// TIA Portal project "SMSS-ENLAB-01-003-1508-012-PLC-B_V13_SP1_1_V17" (V17) (continued)
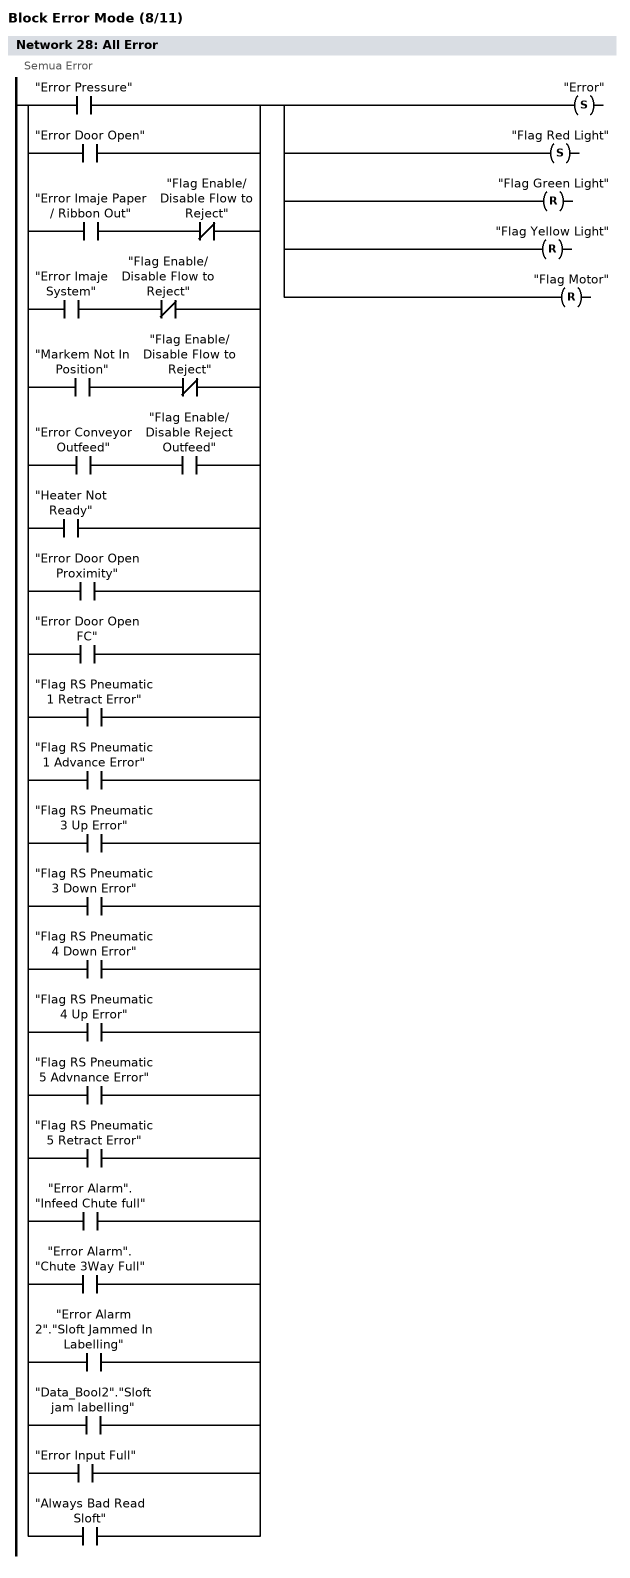
   RUNG wire#powerrail
      Contact( "Error Pressure" )
      wire#w1
      S_Coil( "Error" )
   END_RUNG
   RUNG wire#powerrail
      Contact( "Error Door Open" )
   END_RUNG wire#w1
   RUNG wire#powerrail
      Contact( "Error Imaje Paper / Ribbon Out" )
      I_Contact( "Flag Enable/Disable Flow to Reject" )
   END_RUNG wire#w1
   RUNG wire#powerrail
      Contact( "Error Imaje System" )
      I_Contact( "Flag Enable/Disable Flow to Reject" )
   END_RUNG wire#w1
   RUNG wire#powerrail
      Contact( "Markem Not In Position" )
      I_Contact( "Flag Enable/Disable Flow to Reject" )
   END_RUNG wire#w1
   RUNG wire#powerrail
      Contact( "Error Conveyor Outfeed" )
      Contact( "Flag Enable/Disable Reject Outfeed" )
   END_RUNG wire#w1
   RUNG wire#powerrail
      Contact( "Heater Not Ready" )
   END_RUNG wire#w1
   RUNG wire#powerrail
      Contact( "Error Door Open Proximity" )
   END_RUNG wire#w1
   RUNG wire#powerrail
      Contact( "Error Door Open FC" )
   END_RUNG wire#w1
   RUNG wire#powerrail
      Contact( "Flag RS Pneumatic 1 Retract Error" )
   END_RUNG wire#w1
   RUNG wire#powerrail
      Contact( "Flag RS Pneumatic 1 Advance Error" )
   END_RUNG wire#w1
   RUNG wire#powerrail
      Contact( "Flag RS Pneumatic 3 Up Error" )
   END_RUNG wire#w1
   RUNG wire#powerrail
      Contact( "Flag RS Pneumatic 3 Down Error" )
   END_RUNG wire#w1
   RUNG wire#powerrail
      Contact( "Flag RS Pneumatic 4 Down Error" )
   END_RUNG wire#w1
   RUNG wire#powerrail
      Contact( "Flag RS Pneumatic 4 Up Error" )
   END_RUNG wire#w1
   RUNG wire#powerrail
      Contact( "Flag RS Pneumatic 5 Advnance Error" )
   END_RUNG wire#w1
   RUNG wire#powerrail
      Contact( "Flag RS Pneumatic 5 Retract Error" )
   END_RUNG wire#w1
   RUNG wire#powerrail
      Contact( "Error Alarm"."Infeed Chute full" )
   END_RUNG wire#w1
   RUNG wire#powerrail
      Contact( "Error Alarm"."Chute 3Way Full" )
   END_RUNG wire#w1
   RUNG wire#powerrail
      Contact( "Error Alarm 2"."Sloft Jammed In Labelling" )
   END_RUNG wire#w1
   RUNG wire#powerrail
      Contact( "Data_Bool2"."Sloft jam labelling" )
   END_RUNG wire#w1
   RUNG wire#powerrail
      Contact( "Error Input Full" )
   END_RUNG wire#w1
   RUNG wire#powerrail
      Contact( "Always Bad Read Sloft" )
   END_RUNG wire#w1
   RUNG wire#w1
      S_Coil( "Flag Red Light" )
   END_RUNG
   RUNG wire#w1
      R_Coil( "Flag Green Light" )
   END_RUNG
   RUNG wire#w1
      R_Coil( "Flag Yellow Light" )
   END_RUNG
   RUNG wire#w1
      R_Coil( "Flag Motor" )
   END_RUNG
   // the same network as SCL:
   IF "Error Pressure" OR "Error Door Open" OR ("Error Imaje Paper / Ribbon Out" AND NOT "Flag Enable/Disable Flow to Reject") OR ("Error Imaje System" AND NOT "Flag Enable/Disable Flow to Reject") OR ("Markem Not In Position" AND NOT "Flag Enable/Disable Flow to Reject") OR ("Error Conveyor Outfeed" AND "Flag Enable/Disable Reject Outfeed") OR "Heater Not Ready" OR "Error Door Open Proximity" OR "Error Door Open FC" OR "Flag RS Pneumatic 1 Retract Error" OR "Flag RS Pneumatic 1 Advance Error" OR "Flag RS Pneumatic 3 Up Error" OR "Flag RS Pneumatic 3 Down Error" OR "Flag RS Pneumatic 4 Down Error" OR "Flag RS Pneumatic 4 Up Error" OR "Flag RS Pneumatic 5 Advnance Error" OR "Flag RS Pneumatic 5 Retract Error" OR "Error Alarm"."Infeed Chute full" OR "Error Alarm"."Chute 3Way Full" OR "Error Alarm 2"."Sloft Jammed In Labelling" OR "Data_Bool2"."Sloft jam labelling" OR "Error Input Full" OR "Always Bad Read Sloft" THEN
       "Error" := TRUE;
       "Flag Red Light" := TRUE;
       "Flag Green Light" := FALSE;
       "Flag Yellow Light" := FALSE;
       "Flag Motor" := FALSE;
   END_IF;
END_REGION

REGION Network 29: Reset Error
   // Untuk Reset Semua Error
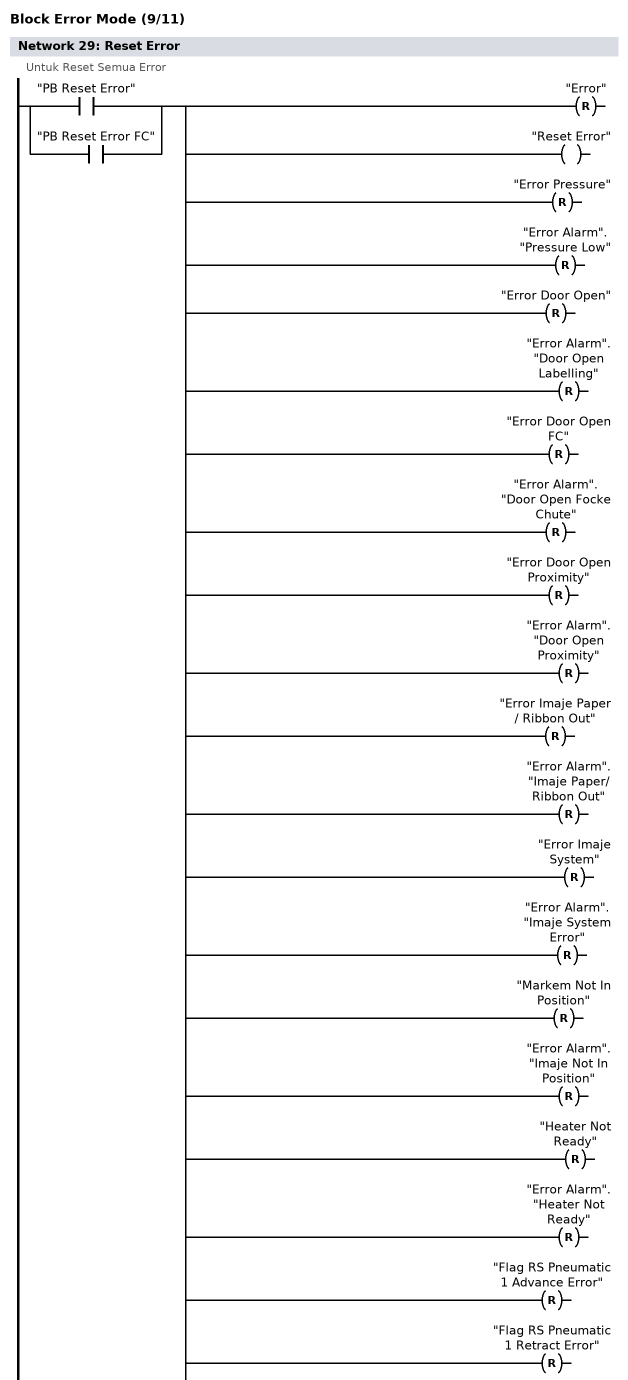
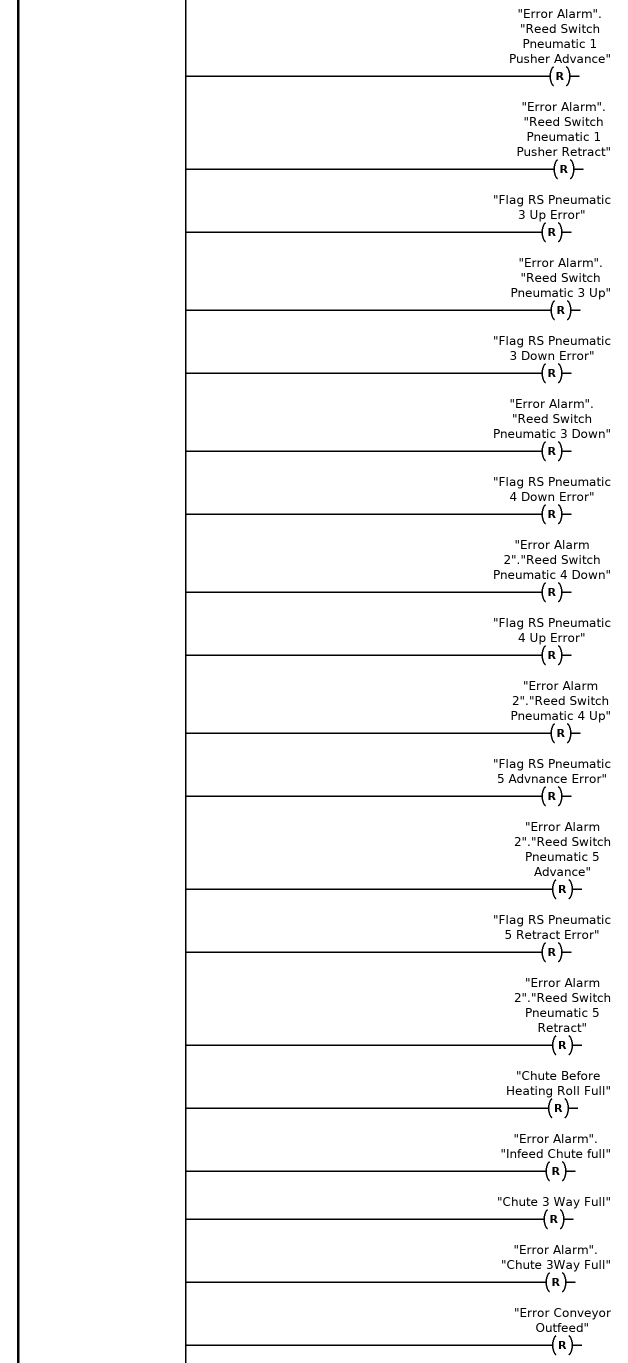
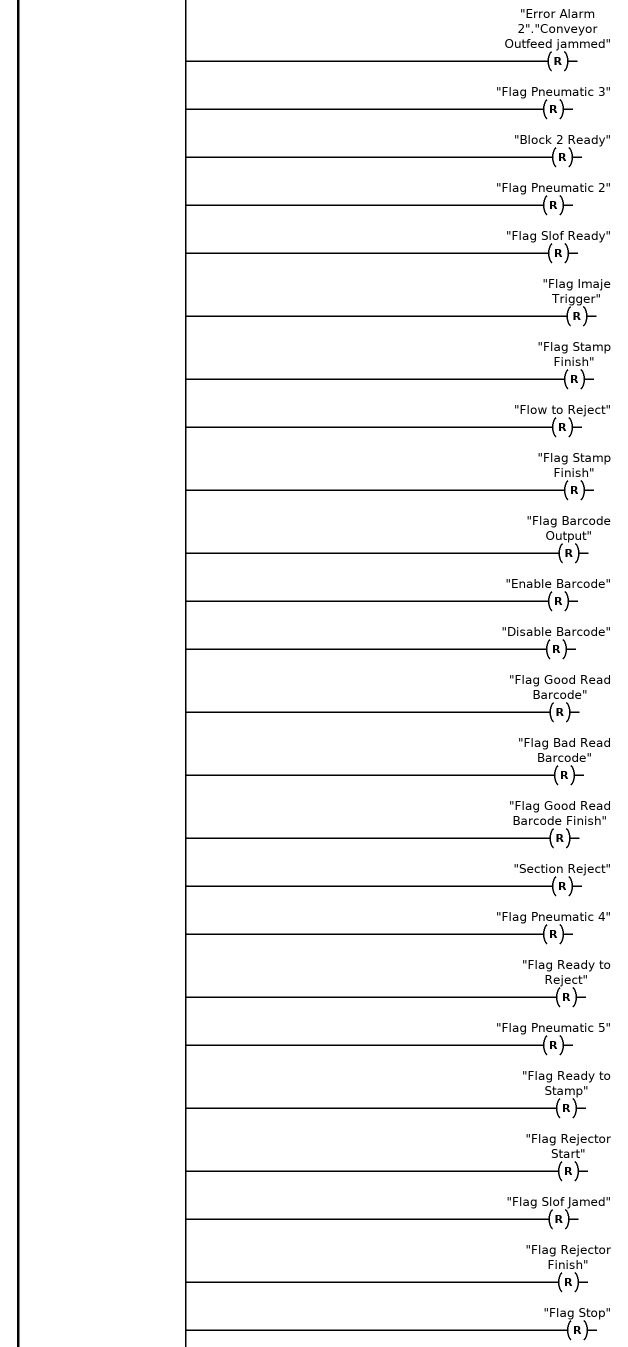
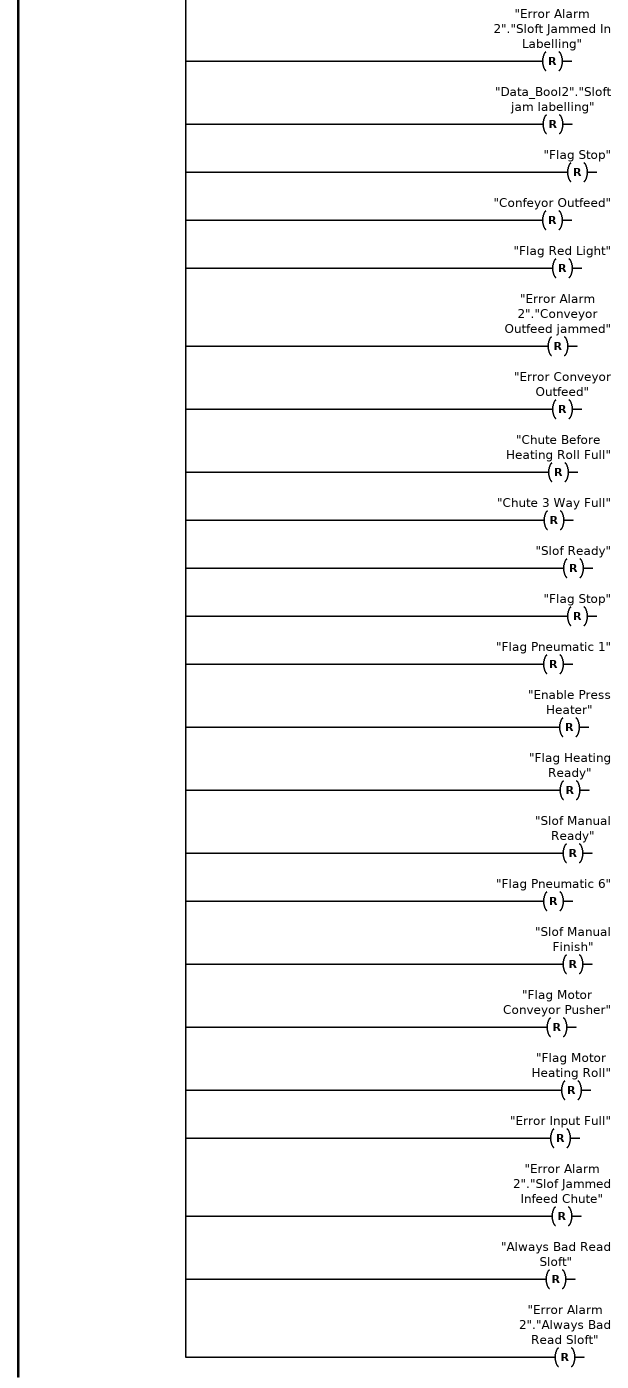
   RUNG wire#powerrail
      Contact( "PB Reset Error" )
      wire#w1
      R_Coil( "Error" )
   END_RUNG
   RUNG wire#powerrail
      Contact( "PB Reset Error FC" )
   END_RUNG wire#w1
   RUNG wire#w1
      Coil( "Reset Error" )
   END_RUNG
   RUNG wire#w1
      R_Coil( "Error Pressure" )
   END_RUNG
   RUNG wire#w1
      R_Coil( "Error Alarm"."Pressure Low" )
   END_RUNG
   RUNG wire#w1
      R_Coil( "Error Door Open" )
   END_RUNG
   RUNG wire#w1
      R_Coil( "Error Alarm"."Door Open Labelling" )
   END_RUNG
   RUNG wire#w1
      R_Coil( "Error Door Open FC" )
   END_RUNG
   RUNG wire#w1
      R_Coil( "Error Alarm"."Door Open Focke Chute" )
   END_RUNG
   RUNG wire#w1
      R_Coil( "Error Door Open Proximity" )
   END_RUNG
   RUNG wire#w1
      R_Coil( "Error Alarm"."Door Open Proximity" )
   END_RUNG
   RUNG wire#w1
      R_Coil( "Error Imaje Paper / Ribbon Out" )
   END_RUNG
   RUNG wire#w1
      R_Coil( "Error Alarm"."Imaje Paper/Ribbon Out" )
   END_RUNG
   RUNG wire#w1
      R_Coil( "Error Imaje System" )
   END_RUNG
   RUNG wire#w1
      R_Coil( "Error Alarm"."Imaje System Error" )
   END_RUNG
   RUNG wire#w1
      R_Coil( "Markem Not In Position" )
   END_RUNG
   RUNG wire#w1
      R_Coil( "Error Alarm"."Imaje Not In Position" )
   END_RUNG
   RUNG wire#w1
      R_Coil( "Heater Not Ready" )
   END_RUNG
   RUNG wire#w1
      R_Coil( "Error Alarm"."Heater Not Ready" )
   END_RUNG
   RUNG wire#w1
      R_Coil( "Flag RS Pneumatic 1 Advance Error" )
   END_RUNG
   RUNG wire#w1
      R_Coil( "Flag RS Pneumatic 1 Retract Error" )
   END_RUNG
   RUNG wire#w1
      R_Coil( "Error Alarm"."Reed Switch Pneumatic 1 Pusher Advance" )
   END_RUNG
   RUNG wire#w1
      R_Coil( "Error Alarm"."Reed Switch Pneumatic 1 Pusher Retract" )
   END_RUNG
   RUNG wire#w1
      R_Coil( "Flag RS Pneumatic 3 Up Error" )
   END_RUNG
   RUNG wire#w1
      R_Coil( "Error Alarm"."Reed Switch Pneumatic 3 Up" )
   END_RUNG
   RUNG wire#w1
      R_Coil( "Flag RS Pneumatic 3 Down Error" )
   END_RUNG
   RUNG wire#w1
      R_Coil( "Error Alarm"."Reed Switch Pneumatic 3 Down" )
   END_RUNG
   RUNG wire#w1
      R_Coil( "Flag RS Pneumatic 4 Down Error" )
   END_RUNG
   RUNG wire#w1
      R_Coil( "Error Alarm 2"."Reed Switch Pneumatic 4 Down" )
   END_RUNG
   RUNG wire#w1
      R_Coil( "Flag RS Pneumatic 4 Up Error" )
   END_RUNG
   RUNG wire#w1
      R_Coil( "Error Alarm 2"."Reed Switch Pneumatic 4 Up" )
   END_RUNG
   RUNG wire#w1
      R_Coil( "Flag RS Pneumatic 5 Advnance Error" )
   END_RUNG
   RUNG wire#w1
      R_Coil( "Error Alarm 2"."Reed Switch Pneumatic 5 Advance" )
   END_RUNG
   RUNG wire#w1
      R_Coil( "Flag RS Pneumatic 5 Retract Error" )
   END_RUNG
   RUNG wire#w1
      R_Coil( "Error Alarm 2"."Reed Switch Pneumatic 5 Retract" )
   END_RUNG
   RUNG wire#w1
      R_Coil( "Chute Before Heating Roll Full" )
   END_RUNG
   RUNG wire#w1
      R_Coil( "Error Alarm"."Infeed Chute full" )
   END_RUNG
   RUNG wire#w1
      R_Coil( "Chute 3 Way Full" )
   END_RUNG
   RUNG wire#w1
      R_Coil( "Error Alarm"."Chute 3Way Full" )
   END_RUNG
   RUNG wire#w1
      R_Coil( "Error Conveyor Outfeed" )
   END_RUNG
   RUNG wire#w1
      R_Coil( "Error Alarm 2"."Conveyor Outfeed jammed" )
   END_RUNG
   RUNG wire#w1
      R_Coil( "Flag Pneumatic 3" )
   END_RUNG
   RUNG wire#w1
      R_Coil( "Block 2 Ready" )
   END_RUNG
   RUNG wire#w1
      R_Coil( "Flag Pneumatic 2" )
   END_RUNG
   RUNG wire#w1
      R_Coil( "Flag Slof Ready" )
   END_RUNG
   RUNG wire#w1
      R_Coil( "Flag Imaje Trigger" )
   END_RUNG
   RUNG wire#w1
      R_Coil( "Flag Stamp Finish" )
   END_RUNG
   RUNG wire#w1
      R_Coil( "Flow to Reject" )
   END_RUNG
   RUNG wire#w1
      R_Coil( "Flag Stamp Finish" )
   END_RUNG
   RUNG wire#w1
      R_Coil( "Flag Barcode Output" )
   END_RUNG
   RUNG wire#w1
      R_Coil( "Enable Barcode" )
   END_RUNG
   RUNG wire#w1
      R_Coil( "Disable Barcode" )
   END_RUNG
   RUNG wire#w1
      R_Coil( "Flag Good Read Barcode" )
   END_RUNG
   RUNG wire#w1
      R_Coil( "Flag Bad Read Barcode" )
   END_RUNG
   RUNG wire#w1
      R_Coil( "Flag Good Read Barcode Finish" )
   END_RUNG
   RUNG wire#w1
      R_Coil( "Section Reject" )
   END_RUNG
   RUNG wire#w1
      R_Coil( "Flag Pneumatic 4" )
   END_RUNG
   RUNG wire#w1
      R_Coil( "Flag Ready to Reject" )
   END_RUNG
   RUNG wire#w1
      R_Coil( "Flag Pneumatic 5" )
   END_RUNG
   RUNG wire#w1
      R_Coil( "Flag Ready to Stamp" )
   END_RUNG
   RUNG wire#w1
      R_Coil( "Flag Rejector Start" )
   END_RUNG
   RUNG wire#w1
      R_Coil( "Flag Slof Jamed" )
   END_RUNG
   RUNG wire#w1
      R_Coil( "Flag Rejector Finish" )
   END_RUNG
   RUNG wire#w1
      R_Coil( "Flag Stop" )
   END_RUNG
   RUNG wire#w1
      R_Coil( "Error Alarm 2"."Sloft Jammed In Labelling" )
   END_RUNG
   RUNG wire#w1
      R_Coil( "Data_Bool2"."Sloft jam labelling" )
   END_RUNG
   RUNG wire#w1
      R_Coil( "Flag Stop" )
   END_RUNG
   RUNG wire#w1
      R_Coil( "Confeyor Outfeed" )
   END_RUNG
   RUNG wire#w1
      R_Coil( "Flag Red Light" )
   END_RUNG
   RUNG wire#w1
      R_Coil( "Error Alarm 2"."Conveyor Outfeed jammed" )
   END_RUNG
   RUNG wire#w1
      R_Coil( "Error Conveyor Outfeed" )
   END_RUNG
   RUNG wire#w1
      R_Coil( "Chute Before Heating Roll Full" )
   END_RUNG
   RUNG wire#w1
      R_Coil( "Chute 3 Way Full" )
   END_RUNG
   RUNG wire#w1
      R_Coil( "Slof Ready" )
   END_RUNG
   RUNG wire#w1
      R_Coil( "Flag Stop" )
   END_RUNG
   RUNG wire#w1
      R_Coil( "Flag Pneumatic 1" )
   END_RUNG
   RUNG wire#w1
      R_Coil( "Enable Press Heater" )
   END_RUNG
   RUNG wire#w1
      R_Coil( "Flag Heating Ready" )
   END_RUNG
   RUNG wire#w1
      R_Coil( "Slof Manual Ready" )
   END_RUNG
   RUNG wire#w1
      R_Coil( "Flag Pneumatic 6" )
   END_RUNG
   RUNG wire#w1
      R_Coil( "Slof Manual Finish" )
   END_RUNG
   RUNG wire#w1
      R_Coil( "Flag Motor Conveyor Pusher" )
   END_RUNG
   RUNG wire#w1
      R_Coil( "Flag Motor Heating Roll" )
   END_RUNG
   RUNG wire#w1
      R_Coil( "Error Input Full" )
   END_RUNG
   RUNG wire#w1
      R_Coil( "Error Alarm 2"."Slof Jammed Infeed Chute" )
   END_RUNG
   RUNG wire#w1
      R_Coil( "Always Bad Read Sloft" )
   END_RUNG
   RUNG wire#w1
      R_Coil( "Error Alarm 2"."Always Bad Read Sloft" )
   END_RUNG
   // the same network as SCL:
   #_w1 := "PB Reset Error" OR "PB Reset Error FC";
   IF #_w1 THEN "Error" := FALSE; END_IF;
   "Reset Error" := #_w1;
   IF #_w1 THEN
       "Error Pressure" := FALSE;
       "Error Alarm"."Pressure Low" := FALSE;
       "Error Door Open" := FALSE;
       "Error Alarm"."Door Open Labelling" := FALSE;
       "Error Door Open FC" := FALSE;
       "Error Alarm"."Door Open Focke Chute" := FALSE;
       "Error Door Open Proximity" := FALSE;
       "Error Alarm"."Door Open Proximity" := FALSE;
       "Error Imaje Paper / Ribbon Out" := FALSE;
       "Error Alarm"."Imaje Paper/Ribbon Out" := FALSE;
       "Error Imaje System" := FALSE;
       "Error Alarm"."Imaje System Error" := FALSE;
       "Markem Not In Position" := FALSE;
       "Error Alarm"."Imaje Not In Position" := FALSE;
       "Heater Not Ready" := FALSE;
       "Error Alarm"."Heater Not Ready" := FALSE;
       "Flag RS Pneumatic 1 Advance Error" := FALSE;
       "Flag RS Pneumatic 1 Retract Error" := FALSE;
       "Error Alarm"."Reed Switch Pneumatic 1 Pusher Advance" := FALSE;
       "Error Alarm"."Reed Switch Pneumatic 1 Pusher Retract" := FALSE;
       "Flag RS Pneumatic 3 Up Error" := FALSE;
       "Error Alarm"."Reed Switch Pneumatic 3 Up" := FALSE;
       "Flag RS Pneumatic 3 Down Error" := FALSE;
       "Error Alarm"."Reed Switch Pneumatic 3 Down" := FALSE;
       "Flag RS Pneumatic 4 Down Error" := FALSE;
       "Error Alarm 2"."Reed Switch Pneumatic 4 Down" := FALSE;
       "Flag RS Pneumatic 4 Up Error" := FALSE;
       "Error Alarm 2"."Reed Switch Pneumatic 4 Up" := FALSE;
       "Flag RS Pneumatic 5 Advnance Error" := FALSE;
       "Error Alarm 2"."Reed Switch Pneumatic 5 Advance" := FALSE;
       "Flag RS Pneumatic 5 Retract Error" := FALSE;
       "Error Alarm 2"."Reed Switch Pneumatic 5 Retract" := FALSE;
       "Chute Before Heating Roll Full" := FALSE;
       "Error Alarm"."Infeed Chute full" := FALSE;
       "Chute 3 Way Full" := FALSE;
       "Error Alarm"."Chute 3Way Full" := FALSE;
       "Error Conveyor Outfeed" := FALSE;
       "Error Alarm 2"."Conveyor Outfeed jammed" := FALSE;
       "Flag Pneumatic 3" := FALSE;
       "Block 2 Ready" := FALSE;
       "Flag Pneumatic 2" := FALSE;
       "Flag Slof Ready" := FALSE;
       "Flag Imaje Trigger" := FALSE;
       "Flag Stamp Finish" := FALSE;
       "Flow to Reject" := FALSE;
       "Flag Stamp Finish" := FALSE;
       "Flag Barcode Output" := FALSE;
       "Enable Barcode" := FALSE;
       "Disable Barcode" := FALSE;
       "Flag Good Read Barcode" := FALSE;
       "Flag Bad Read Barcode" := FALSE;
       "Flag Good Read Barcode Finish" := FALSE;
       "Section Reject" := FALSE;
       "Flag Pneumatic 4" := FALSE;
       "Flag Ready to Reject" := FALSE;
       "Flag Pneumatic 5" := FALSE;
       "Flag Ready to Stamp" := FALSE;
       "Flag Rejector Start" := FALSE;
       "Flag Slof Jamed" := FALSE;
       "Flag Rejector Finish" := FALSE;
       "Flag Stop" := FALSE;
       "Error Alarm 2"."Sloft Jammed In Labelling" := FALSE;
       "Data_Bool2"."Sloft jam labelling" := FALSE;
       "Flag Stop" := FALSE;
       "Confeyor Outfeed" := FALSE;
       "Flag Red Light" := FALSE;
       "Error Alarm 2"."Conveyor Outfeed jammed" := FALSE;
       "Error Conveyor Outfeed" := FALSE;
       "Chute Before Heating Roll Full" := FALSE;
       "Chute 3 Way Full" := FALSE;
       "Slof Ready" := FALSE;
       "Flag Stop" := FALSE;
       "Flag Pneumatic 1" := FALSE;
       "Enable Press Heater" := FALSE;
       "Flag Heating Ready" := FALSE;
       "Slof Manual Ready" := FALSE;
       "Flag Pneumatic 6" := FALSE;
       "Slof Manual Finish" := FALSE;
       "Flag Motor Conveyor Pusher" := FALSE;
       "Flag Motor Heating Roll" := FALSE;
       "Error Input Full" := FALSE;
       "Error Alarm 2"."Slof Jammed Infeed Chute" := FALSE;
       "Always Bad Read Sloft" := FALSE;
       "Error Alarm 2"."Always Bad Read Sloft" := FALSE;
   END_IF;
END_REGION

REGION Network 30: Enable Flow to Reject/Flow To Reject